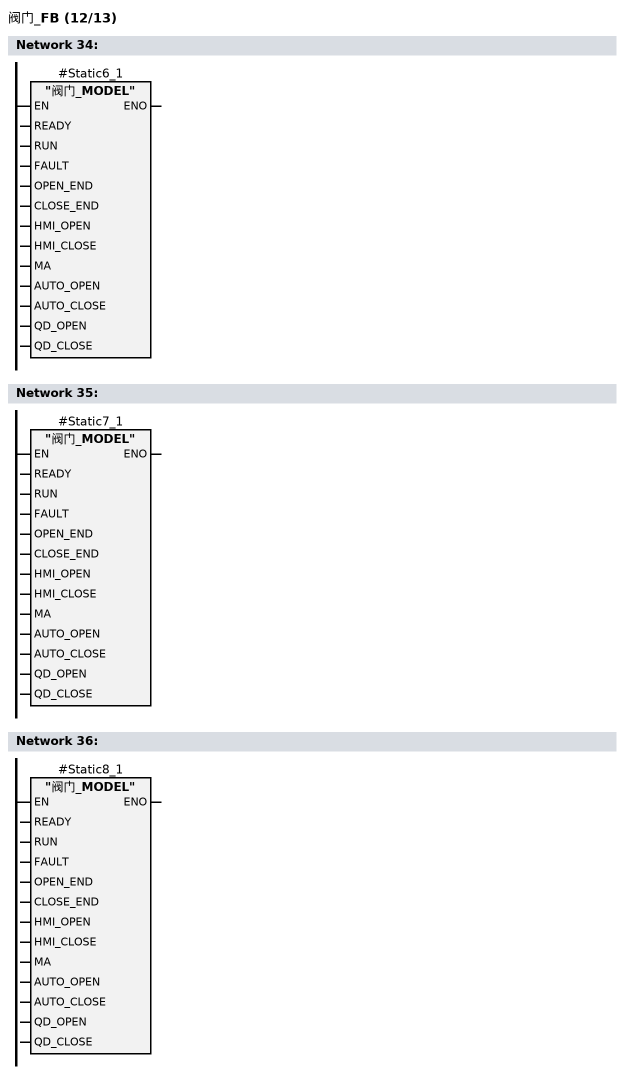
   RUNG wire#powerrail
      #Static6_1(READY :=, RUN :=, FAULT :=, OPEN_END :=, CLOSE_END :=, HMI_OPEN :=, HMI_CLOSE :=, MA :=, AUTO_OPEN :=, AUTO_CLOSE :=, QD_OPEN :=, QD_CLOSE :=)
   END_RUNG
   // the same network as SCL:
   #Static6_1();   // "阀门_MODEL"
END_REGION

REGION Network 35
   RUNG wire#powerrail
      #Static7_1(READY :=, RUN :=, FAULT :=, OPEN_END :=, CLOSE_END :=, HMI_OPEN :=, HMI_CLOSE :=, MA :=, AUTO_OPEN :=, AUTO_CLOSE :=, QD_OPEN :=, QD_CLOSE :=)
   END_RUNG
   // the same network as SCL:
   #Static7_1();   // "阀门_MODEL"
END_REGION

REGION Network 36
   RUNG wire#powerrail
      #Static8_1(READY :=, RUN :=, FAULT :=, OPEN_END :=, CLOSE_END :=, HMI_OPEN :=, HMI_CLOSE :=, MA :=, AUTO_OPEN :=, AUTO_CLOSE :=, QD_OPEN :=, QD_CLOSE :=)
   END_RUNG
   // the same network as SCL:
   #Static8_1();   // "阀门_MODEL"
END_REGION

REGION Network 37
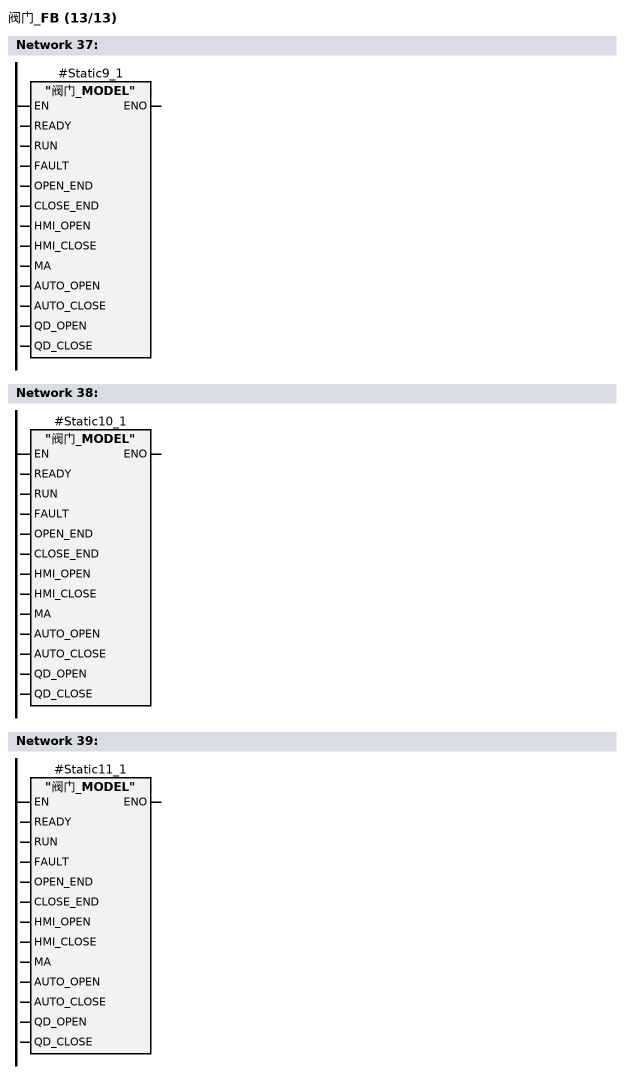
   RUNG wire#powerrail
      #Static9_1(READY :=, RUN :=, FAULT :=, OPEN_END :=, CLOSE_END :=, HMI_OPEN :=, HMI_CLOSE :=, MA :=, AUTO_OPEN :=, AUTO_CLOSE :=, QD_OPEN :=, QD_CLOSE :=)
   END_RUNG
   // the same network as SCL:
   #Static9_1();   // "阀门_MODEL"
END_REGION

REGION Network 38
   RUNG wire#powerrail
      #Static10_1(READY :=, RUN :=, FAULT :=, OPEN_END :=, CLOSE_END :=, HMI_OPEN :=, HMI_CLOSE :=, MA :=, AUTO_OPEN :=, AUTO_CLOSE :=, QD_OPEN :=, QD_CLOSE :=)
   END_RUNG
   // the same network as SCL:
   #Static10_1();   // "阀门_MODEL"
END_REGION

REGION Network 39
   RUNG wire#powerrail
      #Static11_1(READY :=, RUN :=, FAULT :=, OPEN_END :=, CLOSE_END :=, HMI_OPEN :=, HMI_CLOSE :=, MA :=, AUTO_OPEN :=, AUTO_CLOSE :=, QD_OPEN :=, QD_CLOSE :=)
   END_RUNG
   // the same network as SCL:
   #Static11_1();   // "阀门_MODEL"
END_REGION
END_FUNCTION_BLOCK

FUNCTION_BLOCK "引水阀和排气阀FB"   // FB12, LAD
{ S7_Optimized_Access := 'FALSE' }
VERSION : 0.1
   VAR
      "1#炉体循环水泵引水电磁阀" : "引水排气块";
      "1#炉体循环水泵排气电磁阀" : "引水排气块";
      "2#炉体循环水泵引水电磁阀" : "引水排气块";
      "2#炉体循环水泵排气电磁阀" : "引水排气块";
      "3#炉体循环水泵引水电磁阀" : "引水排气块";
      "3#炉体循环水泵排气电磁阀" : "引水排气块";
      "1#电极循环水泵引水电磁阀" : "引水排气块";
      "1#电极循环水泵排气电磁阀" : "引水排气块";
      "2#电极循环水泵引水电磁阀" : "引水排气块";
      "2#电极循环水泵排气电磁阀" : "引水排气块";
      "3#电极循环水泵引水电磁阀" : "引水排气块";
      "3#电极循环水泵排气电磁阀" : "引水排气块";
      "4#电极循环水泵引水电磁阀" : "引水排气块";
      "4#电极循环水泵排气电磁阀" : "引水排气块";
      "1#净环热水泵引水电磁阀" : "引水排气块";
      "1#净环热水泵排气电磁阀" : "引水排气块";
      "2#净环热水泵引水电磁阀" : "引水排气块";
      "2#净环热水泵排气电磁阀" : "引水排气块";
      "3#净环热水泵引水电磁阀" : "引水排气块";
      "3#净环热水泵排气电磁阀" : "引水排气块";
      "4#净环热水泵引水电磁阀" : "引水排气块";
      "4#净环热水泵排气电磁阀" : "引水排气块";
      "5#净环热水泵引水电磁阀" : "引水排气块";
      "5#净环热水泵排气电磁阀" : "引水排气块";
      "1#浊环热水泵引水电磁阀" : "引水排气块";
      "1#浊环热水泵排气电磁阀" : "引水排气块";
      "2#浊环热水泵引水电磁阀" : "引水排气块";
      "2#浊环热水泵排气电磁阀" : "引水排气块";
      "3#浊环热水泵引水电磁阀" : "引水排气块";
      "3#浊环热水泵排气电磁阀" : "引水排气块";
      "4#浊环热水泵引水电磁阀" : "引水排气块";
      "4#浊环热水泵排气电磁阀" : "引水排气块";
      "5#浊环热水泵引水电磁阀" : "引水排气块";
      "5#浊环热水泵排气电磁阀" : "引水排气块";
      "6#浊环热水泵引水电磁阀" : "引水排气块";
      "6#浊环热水泵排气电磁阀" : "引水排气块";
      "7#浊环热水泵引水电磁阀" : "引水排气块";
      "7#浊环热水泵排气电磁阀" : "引水排气块";
      "8#浊环热水泵引水电磁阀" : "引水排气块";
      "8#浊环热水泵排气电磁阀" : "引水排气块";
      "1#冲渣泵引水电磁阀" : "引水排气块";
      "1#冲渣泵排气电磁阀" : "引水排气块";
      "2#冲渣泵引水电磁阀" : "引水排气块";
      "2#冲渣泵排气电磁阀" : "引水排气块";
      "3#冲渣泵引水电磁阀" : "引水排气块";
      "3#冲渣泵排气电磁阀" : "引水排气块";
      "4#冲渣泵引水电磁阀" : "引水排气块";
      "4#冲渣泵排气电磁阀" : "引水排气块";
      "5#冲渣泵引水电磁阀" : "引水排气块";
      "5#冲渣泵排气电磁阀" : "引水排气块";
      "6#冲渣泵引水电磁阀" : "引水排气块";
      "6#冲渣泵排气电磁阀" : "引水排气块";
      "7#冲渣泵引水电磁阀" : "引水排气块";
      "7#冲渣泵排气电磁阀" : "引水排气块";
      "8#冲渣泵引水电磁阀" : "引水排气块";
      "8#冲渣泵排气电磁阀" : "引水排气块";
      "1#柴油泵引水电磁阀" : "引水排气块";
      "1#柴油泵排气电磁阀" : "引水排气块";
      "2#柴油泵引水电磁阀" : "引水排气块";
      "2#柴油泵排气电磁阀" : "引水排气块";
      "1#炉冲渣报警" : "引水排气块";
      "2#炉冲渣报警" : "引水排气块";
      窑冷却泵引水电池阀 : "引水排气块";
      窑冷却泵排气电池阀 : "引水排气块";
      Static9 : "引水排气块";
      Static10 : "引水排气块";
      Static11 : "引水排气块";
      Static12 : "引水排气块";
      Static13 : "引水排气块";
      Static14 : "引水排气块";
      Static15 : "引水排气块";
      Static16 : "引水排气块";
      Static17 : "引水排气块";
      Static18 : "引水排气块";
      Static19 : "引水排气块";
      Static20 : "引水排气块";
      Static21 : "引水排气块";
      Static22 : "引水排气块";
      Static23 : "引水排气块";
      Static24 : "引水排气块";
      Static25 : "引水排气块";
      Static26 : "引水排气块";
      Static27 : "引水排气块";
      Static28 : "引水排气块";
      Static29 : "引水排气块";
      Static30 : "引水排气块";
      Static31 : "引水排气块";
      Static32 : "引水排气块";
      Static33 : "引水排气块";
      Static34 : "引水排气块";
      Static35 : "引水排气块";
      Static36 : "引水排气块";
   END_VAR
BEGIN

REGION Network 1
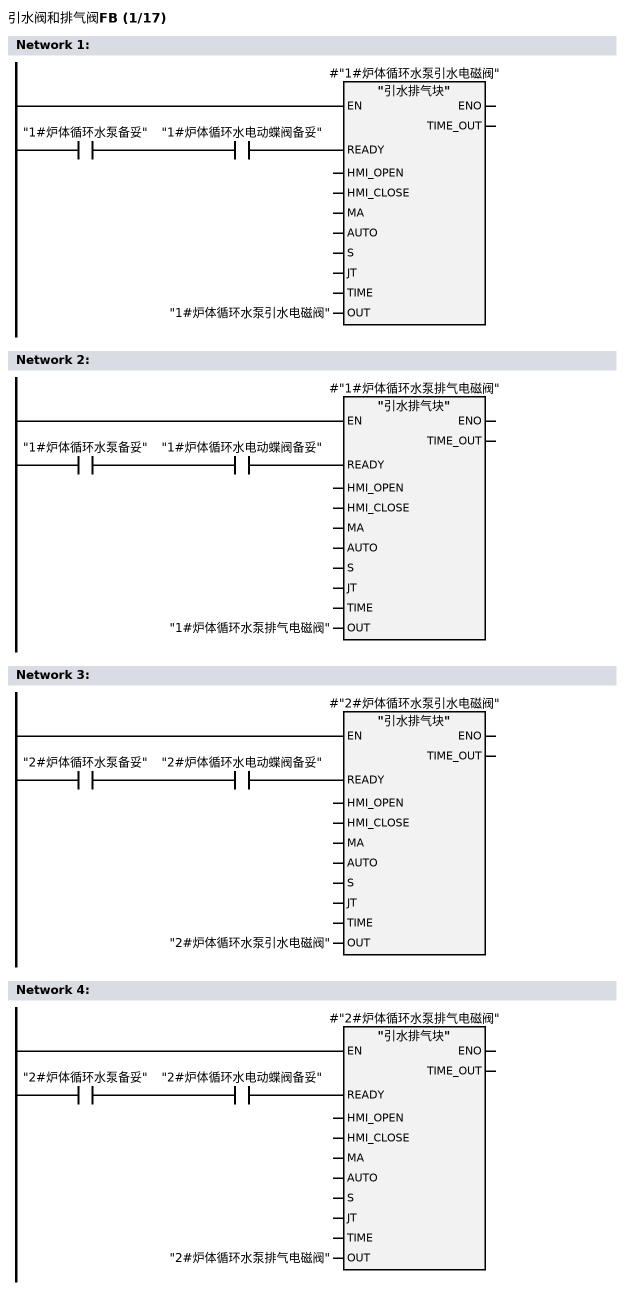
   RUNG wire#powerrail
      #"1#炉体循环水泵引水电磁阀"(READY := wire#w1, HMI_OPEN :=, HMI_CLOSE :=, MA :=, AUTO :=, S :=, JT :=, "TIME" :=, OUT := "1#炉体循环水泵引水电磁阀", TIME_OUT =>)
   END_RUNG
   RUNG wire#powerrail
      Contact( "1#炉体循环水泵备妥" )
      Contact( "1#炉体循环水电动蝶阀备妥" )
   END_RUNG wire#w1
   // the same network as SCL:
   #"1#炉体循环水泵引水电磁阀"(READY := "1#炉体循环水泵备妥" AND "1#炉体循环水电动蝶阀备妥", OUT := "1#炉体循环水泵引水电磁阀");   // "引水排气块"
END_REGION

REGION Network 2
   RUNG wire#powerrail
      #"1#炉体循环水泵排气电磁阀"(READY := wire#w1, HMI_OPEN :=, HMI_CLOSE :=, MA :=, AUTO :=, S :=, JT :=, "TIME" :=, OUT := "1#炉体循环水泵排气电磁阀", TIME_OUT =>)
   END_RUNG
   RUNG wire#powerrail
      Contact( "1#炉体循环水泵备妥" )
      Contact( "1#炉体循环水电动蝶阀备妥" )
   END_RUNG wire#w1
   // the same network as SCL:
   #"1#炉体循环水泵排气电磁阀"(READY := "1#炉体循环水泵备妥" AND "1#炉体循环水电动蝶阀备妥", OUT := "1#炉体循环水泵排气电磁阀");   // "引水排气块"
END_REGION

REGION Network 3
   RUNG wire#powerrail
      #"2#炉体循环水泵引水电磁阀"(READY := wire#w1, HMI_OPEN :=, HMI_CLOSE :=, MA :=, AUTO :=, S :=, JT :=, "TIME" :=, OUT := "2#炉体循环水泵引水电磁阀", TIME_OUT =>)
   END_RUNG
   RUNG wire#powerrail
      Contact( "2#炉体循环水泵备妥" )
      Contact( "2#炉体循环水电动蝶阀备妥" )
   END_RUNG wire#w1
   // the same network as SCL:
   #"2#炉体循环水泵引水电磁阀"(READY := "2#炉体循环水泵备妥" AND "2#炉体循环水电动蝶阀备妥", OUT := "2#炉体循环水泵引水电磁阀");   // "引水排气块"
END_REGION

REGION Network 4
   RUNG wire#powerrail
      #"2#炉体循环水泵排气电磁阀"(READY := wire#w1, HMI_OPEN :=, HMI_CLOSE :=, MA :=, AUTO :=, S :=, JT :=, "TIME" :=, OUT := "2#炉体循环水泵排气电磁阀", TIME_OUT =>)
   END_RUNG
   RUNG wire#powerrail
      Contact( "2#炉体循环水泵备妥" )
      Contact( "2#炉体循环水电动蝶阀备妥" )
   END_RUNG wire#w1
   // the same network as SCL:
   #"2#炉体循环水泵排气电磁阀"(READY := "2#炉体循环水泵备妥" AND "2#炉体循环水电动蝶阀备妥", OUT := "2#炉体循环水泵排气电磁阀");   // "引水排气块"
END_REGION

REGION Network 5
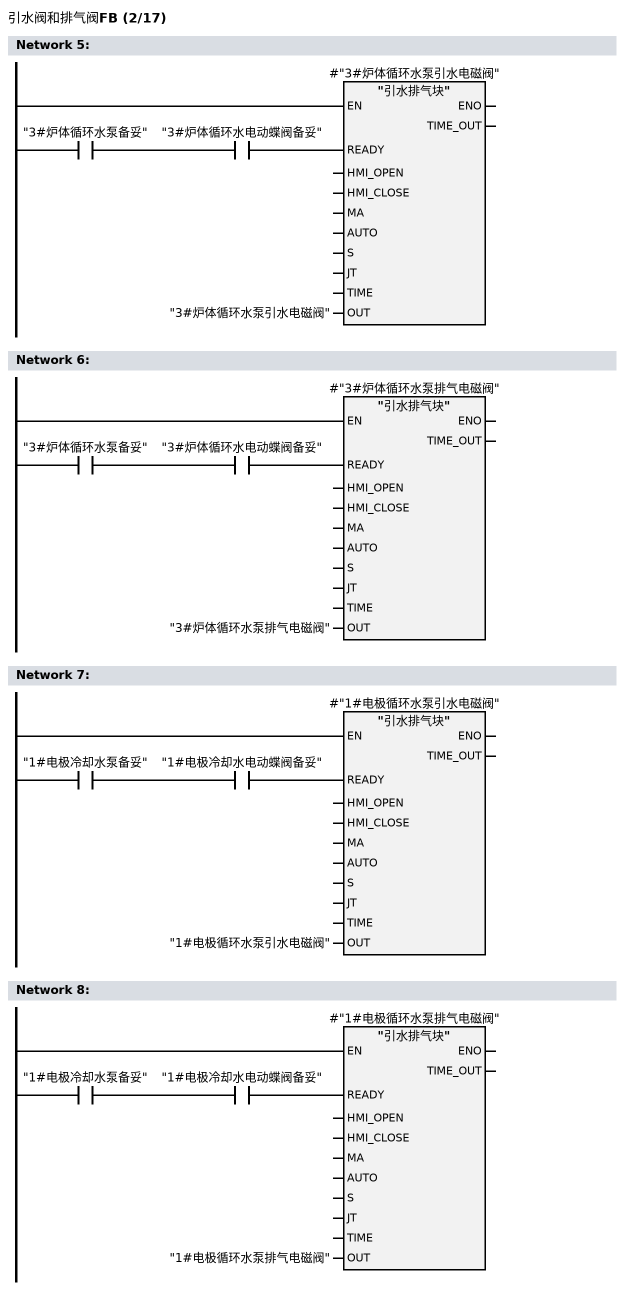
   RUNG wire#powerrail
      #"3#炉体循环水泵引水电磁阀"(READY := wire#w1, HMI_OPEN :=, HMI_CLOSE :=, MA :=, AUTO :=, S :=, JT :=, "TIME" :=, OUT := "3#炉体循环水泵引水电磁阀", TIME_OUT =>)
   END_RUNG
   RUNG wire#powerrail
      Contact( "3#炉体循环水泵备妥" )
      Contact( "3#炉体循环水电动蝶阀备妥" )
   END_RUNG wire#w1
   // the same network as SCL:
   #"3#炉体循环水泵引水电磁阀"(READY := "3#炉体循环水泵备妥" AND "3#炉体循环水电动蝶阀备妥", OUT := "3#炉体循环水泵引水电磁阀");   // "引水排气块"
END_REGION

REGION Network 6
   RUNG wire#powerrail
      #"3#炉体循环水泵排气电磁阀"(READY := wire#w1, HMI_OPEN :=, HMI_CLOSE :=, MA :=, AUTO :=, S :=, JT :=, "TIME" :=, OUT := "3#炉体循环水泵排气电磁阀", TIME_OUT =>)
   END_RUNG
   RUNG wire#powerrail
      Contact( "3#炉体循环水泵备妥" )
      Contact( "3#炉体循环水电动蝶阀备妥" )
   END_RUNG wire#w1
   // the same network as SCL:
   #"3#炉体循环水泵排气电磁阀"(READY := "3#炉体循环水泵备妥" AND "3#炉体循环水电动蝶阀备妥", OUT := "3#炉体循环水泵排气电磁阀");   // "引水排气块"
END_REGION

REGION Network 7
   RUNG wire#powerrail
      #"1#电极循环水泵引水电磁阀"(READY := wire#w1, HMI_OPEN :=, HMI_CLOSE :=, MA :=, AUTO :=, S :=, JT :=, "TIME" :=, OUT := "1#电极循环水泵引水电磁阀", TIME_OUT =>)
   END_RUNG
   RUNG wire#powerrail
      Contact( "1#电极冷却水泵备妥" )
      Contact( "1#电极冷却水电动蝶阀备妥" )
   END_RUNG wire#w1
   // the same network as SCL:
   #"1#电极循环水泵引水电磁阀"(READY := "1#电极冷却水泵备妥" AND "1#电极冷却水电动蝶阀备妥", OUT := "1#电极循环水泵引水电磁阀");   // "引水排气块"
END_REGION

REGION Network 8
   RUNG wire#powerrail
      #"1#电极循环水泵排气电磁阀"(READY := wire#w1, HMI_OPEN :=, HMI_CLOSE :=, MA :=, AUTO :=, S :=, JT :=, "TIME" :=, OUT := "1#电极循环水泵排气电磁阀", TIME_OUT =>)
   END_RUNG
   RUNG wire#powerrail
      Contact( "1#电极冷却水泵备妥" )
      Contact( "1#电极冷却水电动蝶阀备妥" )
   END_RUNG wire#w1
   // the same network as SCL:
   #"1#电极循环水泵排气电磁阀"(READY := "1#电极冷却水泵备妥" AND "1#电极冷却水电动蝶阀备妥", OUT := "1#电极循环水泵排气电磁阀");   // "引水排气块"
END_REGION

REGION Network 9
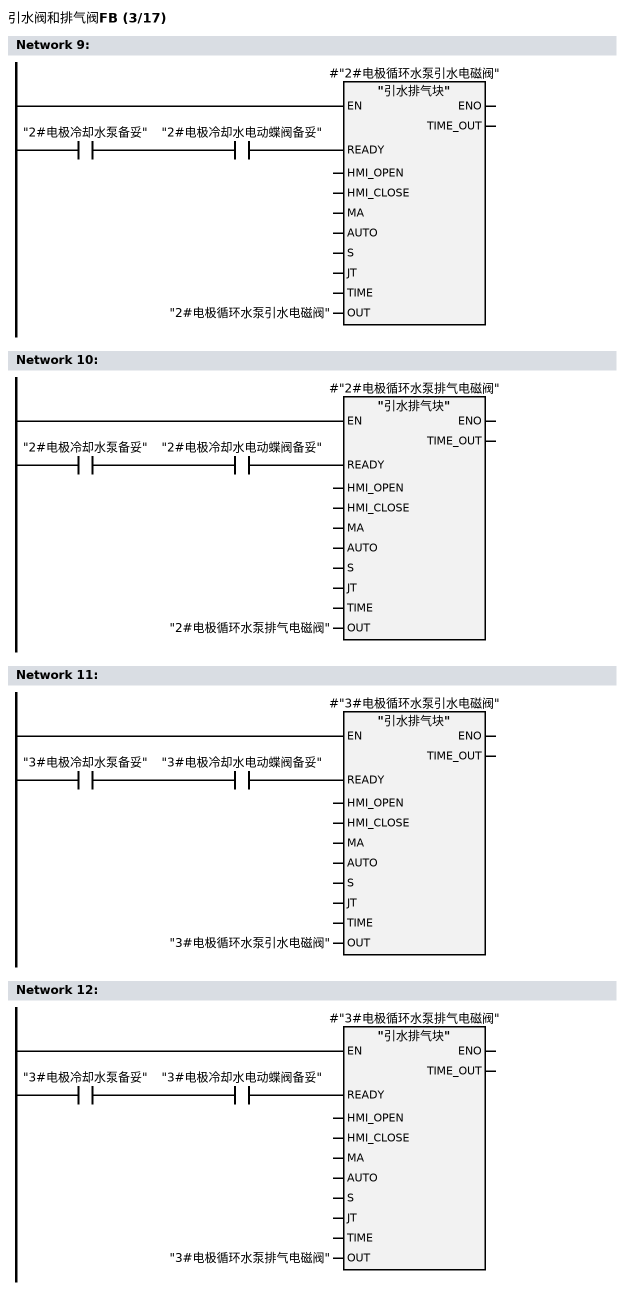
   RUNG wire#powerrail
      #"2#电极循环水泵引水电磁阀"(READY := wire#w1, HMI_OPEN :=, HMI_CLOSE :=, MA :=, AUTO :=, S :=, JT :=, "TIME" :=, OUT := "2#电极循环水泵引水电磁阀", TIME_OUT =>)
   END_RUNG
   RUNG wire#powerrail
      Contact( "2#电极冷却水泵备妥" )
      Contact( "2#电极冷却水电动蝶阀备妥" )
   END_RUNG wire#w1
   // the same network as SCL:
   #"2#电极循环水泵引水电磁阀"(READY := "2#电极冷却水泵备妥" AND "2#电极冷却水电动蝶阀备妥", OUT := "2#电极循环水泵引水电磁阀");   // "引水排气块"
END_REGION

REGION Network 10
   RUNG wire#powerrail
      #"2#电极循环水泵排气电磁阀"(READY := wire#w1, HMI_OPEN :=, HMI_CLOSE :=, MA :=, AUTO :=, S :=, JT :=, "TIME" :=, OUT := "2#电极循环水泵排气电磁阀", TIME_OUT =>)
   END_RUNG
   RUNG wire#powerrail
      Contact( "2#电极冷却水泵备妥" )
      Contact( "2#电极冷却水电动蝶阀备妥" )
   END_RUNG wire#w1
   // the same network as SCL:
   #"2#电极循环水泵排气电磁阀"(READY := "2#电极冷却水泵备妥" AND "2#电极冷却水电动蝶阀备妥", OUT := "2#电极循环水泵排气电磁阀");   // "引水排气块"
END_REGION

REGION Network 11
   RUNG wire#powerrail
      #"3#电极循环水泵引水电磁阀"(READY := wire#w1, HMI_OPEN :=, HMI_CLOSE :=, MA :=, AUTO :=, S :=, JT :=, "TIME" :=, OUT := "3#电极循环水泵引水电磁阀", TIME_OUT =>)
   END_RUNG
   RUNG wire#powerrail
      Contact( "3#电极冷却水泵备妥" )
      Contact( "3#电极冷却水电动蝶阀备妥" )
   END_RUNG wire#w1
   // the same network as SCL:
   #"3#电极循环水泵引水电磁阀"(READY := "3#电极冷却水泵备妥" AND "3#电极冷却水电动蝶阀备妥", OUT := "3#电极循环水泵引水电磁阀");   // "引水排气块"
END_REGION

REGION Network 12
   RUNG wire#powerrail
      #"3#电极循环水泵排气电磁阀"(READY := wire#w1, HMI_OPEN :=, HMI_CLOSE :=, MA :=, AUTO :=, S :=, JT :=, "TIME" :=, OUT := "3#电极循环水泵排气电磁阀", TIME_OUT =>)
   END_RUNG
   RUNG wire#powerrail
      Contact( "3#电极冷却水泵备妥" )
      Contact( "3#电极冷却水电动蝶阀备妥" )
   END_RUNG wire#w1
   // the same network as SCL:
   #"3#电极循环水泵排气电磁阀"(READY := "3#电极冷却水泵备妥" AND "3#电极冷却水电动蝶阀备妥", OUT := "3#电极循环水泵排气电磁阀");   // "引水排气块"
END_REGION

REGION Network 13
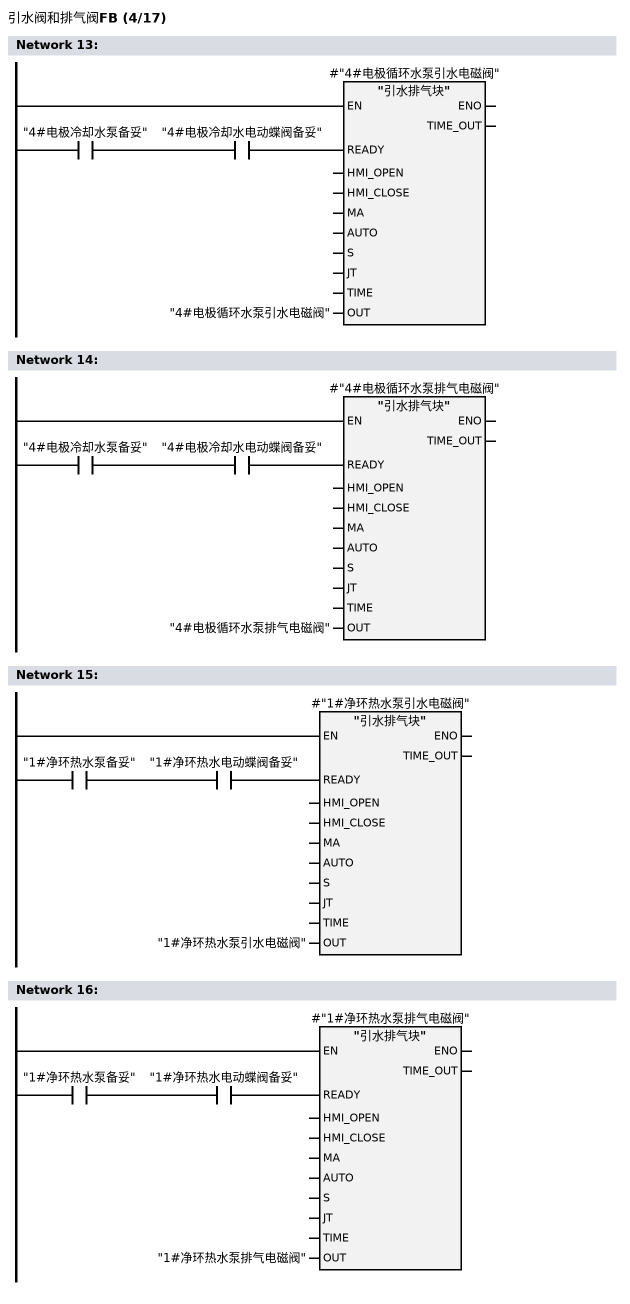
   RUNG wire#powerrail
      #"4#电极循环水泵引水电磁阀"(READY := wire#w1, HMI_OPEN :=, HMI_CLOSE :=, MA :=, AUTO :=, S :=, JT :=, "TIME" :=, OUT := "4#电极循环水泵引水电磁阀", TIME_OUT =>)
   END_RUNG
   RUNG wire#powerrail
      Contact( "4#电极冷却水泵备妥" )
      Contact( "4#电极冷却水电动蝶阀备妥" )
   END_RUNG wire#w1
   // the same network as SCL:
   #"4#电极循环水泵引水电磁阀"(READY := "4#电极冷却水泵备妥" AND "4#电极冷却水电动蝶阀备妥", OUT := "4#电极循环水泵引水电磁阀");   // "引水排气块"
END_REGION

REGION Network 14
   RUNG wire#powerrail
      #"4#电极循环水泵排气电磁阀"(READY := wire#w1, HMI_OPEN :=, HMI_CLOSE :=, MA :=, AUTO :=, S :=, JT :=, "TIME" :=, OUT := "4#电极循环水泵排气电磁阀", TIME_OUT =>)
   END_RUNG
   RUNG wire#powerrail
      Contact( "4#电极冷却水泵备妥" )
      Contact( "4#电极冷却水电动蝶阀备妥" )
   END_RUNG wire#w1
   // the same network as SCL:
   #"4#电极循环水泵排气电磁阀"(READY := "4#电极冷却水泵备妥" AND "4#电极冷却水电动蝶阀备妥", OUT := "4#电极循环水泵排气电磁阀");   // "引水排气块"
END_REGION

REGION Network 15
   RUNG wire#powerrail
      #"1#净环热水泵引水电磁阀"(READY := wire#w1, HMI_OPEN :=, HMI_CLOSE :=, MA :=, AUTO :=, S :=, JT :=, "TIME" :=, OUT := "1#净环热水泵引水电磁阀", TIME_OUT =>)
   END_RUNG
   RUNG wire#powerrail
      Contact( "1#净环热水泵备妥" )
      Contact( "1#净环热水电动蝶阀备妥" )
   END_RUNG wire#w1
   // the same network as SCL:
   #"1#净环热水泵引水电磁阀"(READY := "1#净环热水泵备妥" AND "1#净环热水电动蝶阀备妥", OUT := "1#净环热水泵引水电磁阀");   // "引水排气块"
END_REGION

REGION Network 16
   RUNG wire#powerrail
      #"1#净环热水泵排气电磁阀"(READY := wire#w1, HMI_OPEN :=, HMI_CLOSE :=, MA :=, AUTO :=, S :=, JT :=, "TIME" :=, OUT := "1#净环热水泵排气电磁阀", TIME_OUT =>)
   END_RUNG
   RUNG wire#powerrail
      Contact( "1#净环热水泵备妥" )
      Contact( "1#净环热水电动蝶阀备妥" )
   END_RUNG wire#w1
   // the same network as SCL:
   #"1#净环热水泵排气电磁阀"(READY := "1#净环热水泵备妥" AND "1#净环热水电动蝶阀备妥", OUT := "1#净环热水泵排气电磁阀");   // "引水排气块"
END_REGION

REGION Network 17
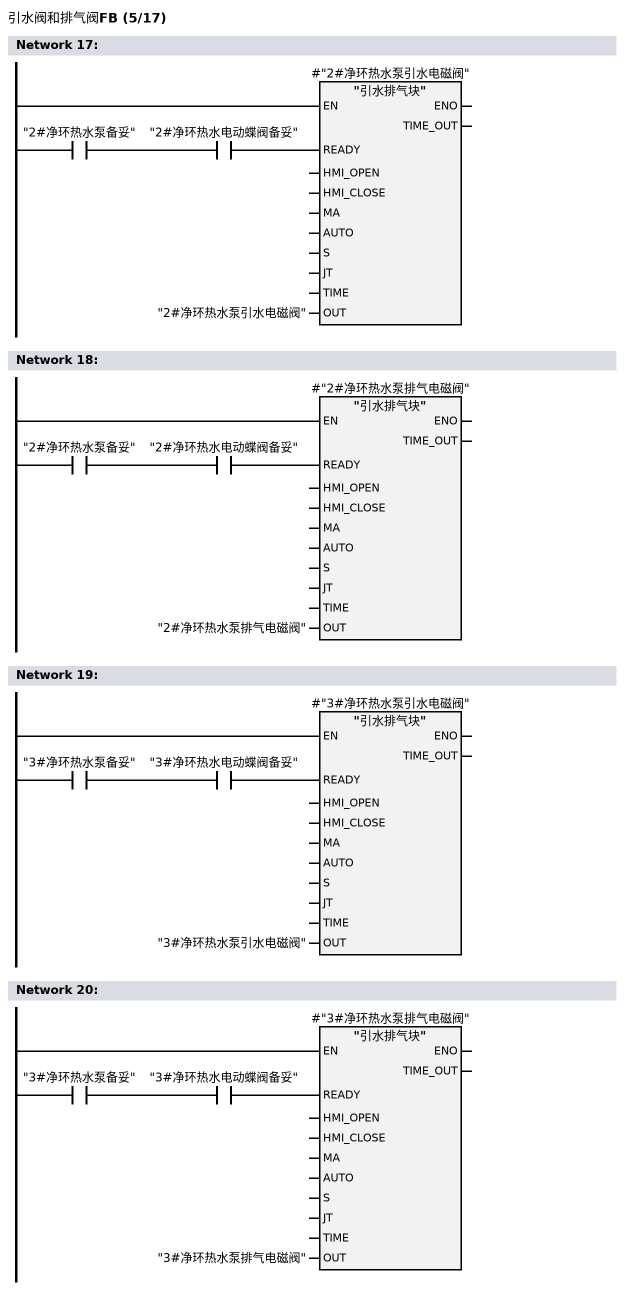
   RUNG wire#powerrail
      #"2#净环热水泵引水电磁阀"(READY := wire#w1, HMI_OPEN :=, HMI_CLOSE :=, MA :=, AUTO :=, S :=, JT :=, "TIME" :=, OUT := "2#净环热水泵引水电磁阀", TIME_OUT =>)
   END_RUNG
   RUNG wire#powerrail
      Contact( "2#净环热水泵备妥" )
      Contact( "2#净环热水电动蝶阀备妥" )
   END_RUNG wire#w1
   // the same network as SCL:
   #"2#净环热水泵引水电磁阀"(READY := "2#净环热水泵备妥" AND "2#净环热水电动蝶阀备妥", OUT := "2#净环热水泵引水电磁阀");   // "引水排气块"
END_REGION

REGION Network 18
   RUNG wire#powerrail
      #"2#净环热水泵排气电磁阀"(READY := wire#w1, HMI_OPEN :=, HMI_CLOSE :=, MA :=, AUTO :=, S :=, JT :=, "TIME" :=, OUT := "2#净环热水泵排气电磁阀", TIME_OUT =>)
   END_RUNG
   RUNG wire#powerrail
      Contact( "2#净环热水泵备妥" )
      Contact( "2#净环热水电动蝶阀备妥" )
   END_RUNG wire#w1
   // the same network as SCL:
   #"2#净环热水泵排气电磁阀"(READY := "2#净环热水泵备妥" AND "2#净环热水电动蝶阀备妥", OUT := "2#净环热水泵排气电磁阀");   // "引水排气块"
END_REGION

REGION Network 19
   RUNG wire#powerrail
      #"3#净环热水泵引水电磁阀"(READY := wire#w1, HMI_OPEN :=, HMI_CLOSE :=, MA :=, AUTO :=, S :=, JT :=, "TIME" :=, OUT := "3#净环热水泵引水电磁阀", TIME_OUT =>)
   END_RUNG
   RUNG wire#powerrail
      Contact( "3#净环热水泵备妥" )
      Contact( "3#净环热水电动蝶阀备妥" )
   END_RUNG wire#w1
   // the same network as SCL:
   #"3#净环热水泵引水电磁阀"(READY := "3#净环热水泵备妥" AND "3#净环热水电动蝶阀备妥", OUT := "3#净环热水泵引水电磁阀");   // "引水排气块"
END_REGION

REGION Network 20
   RUNG wire#powerrail
      #"3#净环热水泵排气电磁阀"(READY := wire#w1, HMI_OPEN :=, HMI_CLOSE :=, MA :=, AUTO :=, S :=, JT :=, "TIME" :=, OUT := "3#净环热水泵排气电磁阀", TIME_OUT =>)
   END_RUNG
   RUNG wire#powerrail
      Contact( "3#净环热水泵备妥" )
      Contact( "3#净环热水电动蝶阀备妥" )
   END_RUNG wire#w1
   // the same network as SCL:
   #"3#净环热水泵排气电磁阀"(READY := "3#净环热水泵备妥" AND "3#净环热水电动蝶阀备妥", OUT := "3#净环热水泵排气电磁阀");   // "引水排气块"
END_REGION

REGION Network 21
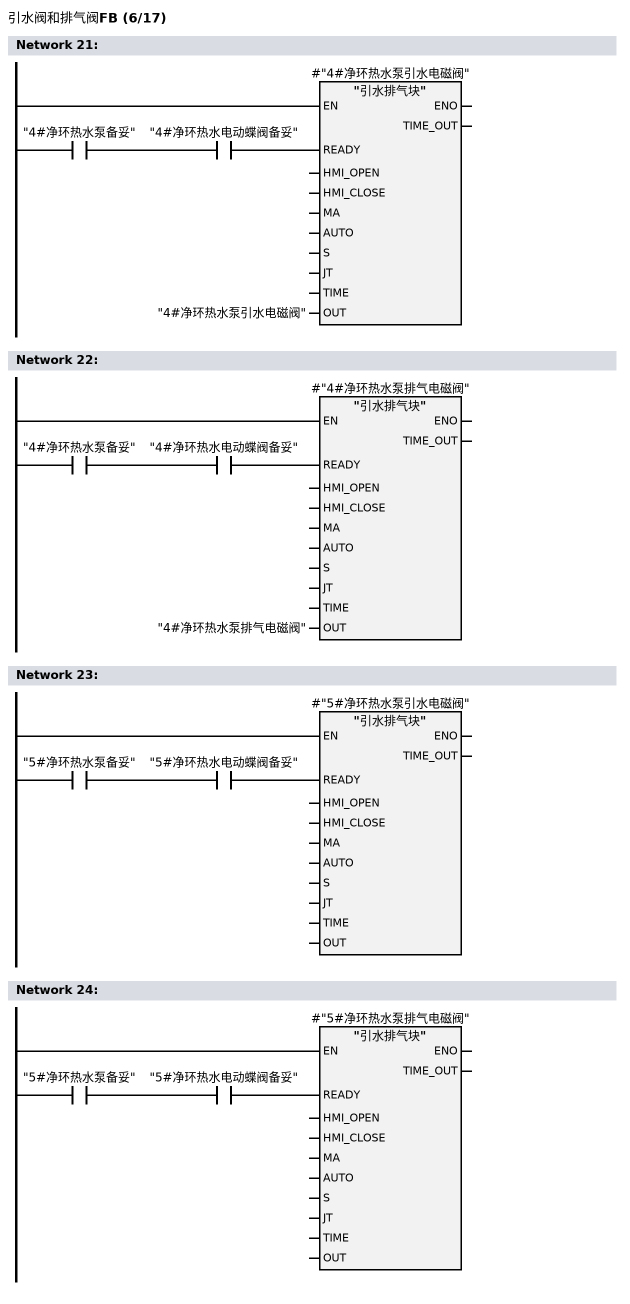
   RUNG wire#powerrail
      #"4#净环热水泵引水电磁阀"(READY := wire#w1, HMI_OPEN :=, HMI_CLOSE :=, MA :=, AUTO :=, S :=, JT :=, "TIME" :=, OUT := "4#净环热水泵引水电磁阀", TIME_OUT =>)
   END_RUNG
   RUNG wire#powerrail
      Contact( "4#净环热水泵备妥" )
      Contact( "4#净环热水电动蝶阀备妥" )
   END_RUNG wire#w1
   // the same network as SCL:
   #"4#净环热水泵引水电磁阀"(READY := "4#净环热水泵备妥" AND "4#净环热水电动蝶阀备妥", OUT := "4#净环热水泵引水电磁阀");   // "引水排气块"
END_REGION

REGION Network 22
   RUNG wire#powerrail
      #"4#净环热水泵排气电磁阀"(READY := wire#w1, HMI_OPEN :=, HMI_CLOSE :=, MA :=, AUTO :=, S :=, JT :=, "TIME" :=, OUT := "4#净环热水泵排气电磁阀", TIME_OUT =>)
   END_RUNG
   RUNG wire#powerrail
      Contact( "4#净环热水泵备妥" )
      Contact( "4#净环热水电动蝶阀备妥" )
   END_RUNG wire#w1
   // the same network as SCL:
   #"4#净环热水泵排气电磁阀"(READY := "4#净环热水泵备妥" AND "4#净环热水电动蝶阀备妥", OUT := "4#净环热水泵排气电磁阀");   // "引水排气块"
END_REGION

REGION Network 23
   RUNG wire#powerrail
      #"5#净环热水泵引水电磁阀"(READY := wire#w1, HMI_OPEN :=, HMI_CLOSE :=, MA :=, AUTO :=, S :=, JT :=, "TIME" :=, OUT :=, TIME_OUT =>)
   END_RUNG
   RUNG wire#powerrail
      Contact( "5#净环热水泵备妥" )
      Contact( "5#净环热水电动蝶阀备妥" )
   END_RUNG wire#w1
   // the same network as SCL:
   #"5#净环热水泵引水电磁阀"(READY := "5#净环热水泵备妥" AND "5#净环热水电动蝶阀备妥");   // "引水排气块"
END_REGION

REGION Network 24
   RUNG wire#powerrail
      #"5#净环热水泵排气电磁阀"(READY := wire#w1, HMI_OPEN :=, HMI_CLOSE :=, MA :=, AUTO :=, S :=, JT :=, "TIME" :=, OUT :=, TIME_OUT =>)
   END_RUNG
   RUNG wire#powerrail
      Contact( "5#净环热水泵备妥" )
      Contact( "5#净环热水电动蝶阀备妥" )
   END_RUNG wire#w1
   // the same network as SCL:
   #"5#净环热水泵排气电磁阀"(READY := "5#净环热水泵备妥" AND "5#净环热水电动蝶阀备妥");   // "引水排气块"
END_REGION

REGION Network 25
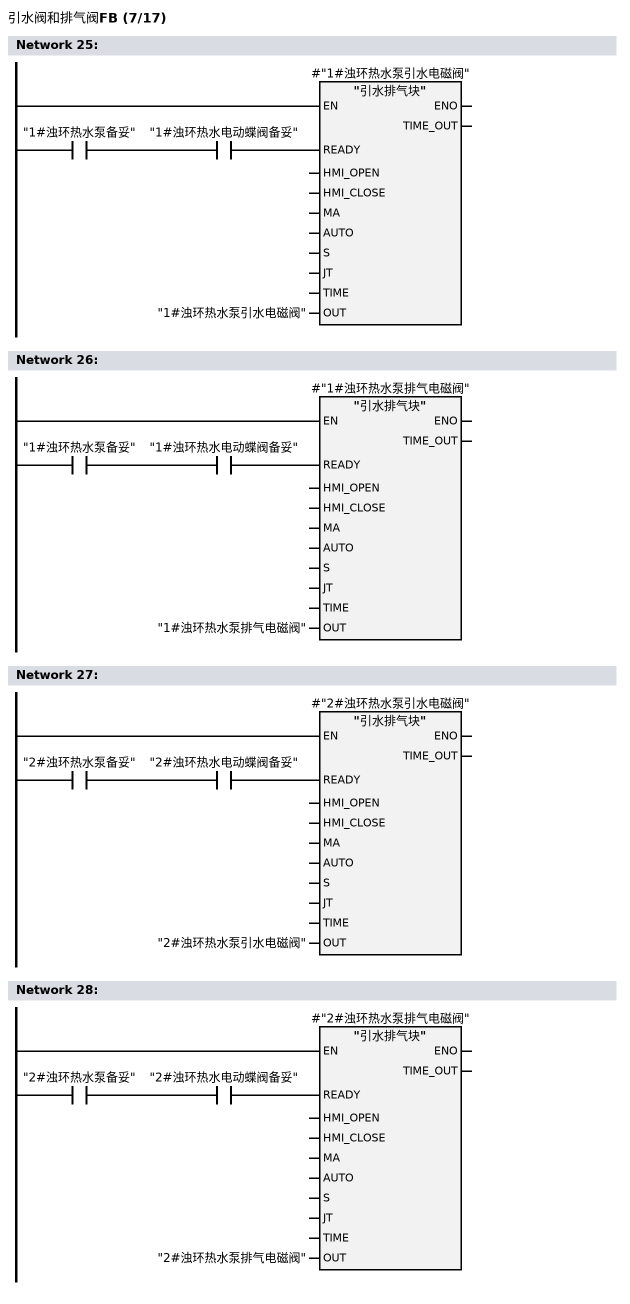
   RUNG wire#powerrail
      #"1#浊环热水泵引水电磁阀"(READY := wire#w1, HMI_OPEN :=, HMI_CLOSE :=, MA :=, AUTO :=, S :=, JT :=, "TIME" :=, OUT := "1#浊环热水泵引水电磁阀", TIME_OUT =>)
   END_RUNG
   RUNG wire#powerrail
      Contact( "1#浊环热水泵备妥" )
      Contact( "1#浊环热水电动蝶阀备妥" )
   END_RUNG wire#w1
   // the same network as SCL:
   #"1#浊环热水泵引水电磁阀"(READY := "1#浊环热水泵备妥" AND "1#浊环热水电动蝶阀备妥", OUT := "1#浊环热水泵引水电磁阀");   // "引水排气块"
END_REGION

REGION Network 26
   RUNG wire#powerrail
      #"1#浊环热水泵排气电磁阀"(READY := wire#w1, HMI_OPEN :=, HMI_CLOSE :=, MA :=, AUTO :=, S :=, JT :=, "TIME" :=, OUT := "1#浊环热水泵排气电磁阀", TIME_OUT =>)
   END_RUNG
   RUNG wire#powerrail
      Contact( "1#浊环热水泵备妥" )
      Contact( "1#浊环热水电动蝶阀备妥" )
   END_RUNG wire#w1
   // the same network as SCL:
   #"1#浊环热水泵排气电磁阀"(READY := "1#浊环热水泵备妥" AND "1#浊环热水电动蝶阀备妥", OUT := "1#浊环热水泵排气电磁阀");   // "引水排气块"
END_REGION

REGION Network 27
   RUNG wire#powerrail
      #"2#浊环热水泵引水电磁阀"(READY := wire#w1, HMI_OPEN :=, HMI_CLOSE :=, MA :=, AUTO :=, S :=, JT :=, "TIME" :=, OUT := "2#浊环热水泵引水电磁阀", TIME_OUT =>)
   END_RUNG
   RUNG wire#powerrail
      Contact( "2#浊环热水泵备妥" )
      Contact( "2#浊环热水电动蝶阀备妥" )
   END_RUNG wire#w1
   // the same network as SCL:
   #"2#浊环热水泵引水电磁阀"(READY := "2#浊环热水泵备妥" AND "2#浊环热水电动蝶阀备妥", OUT := "2#浊环热水泵引水电磁阀");   // "引水排气块"
END_REGION

REGION Network 28
   RUNG wire#powerrail
      #"2#浊环热水泵排气电磁阀"(READY := wire#w1, HMI_OPEN :=, HMI_CLOSE :=, MA :=, AUTO :=, S :=, JT :=, "TIME" :=, OUT := "2#浊环热水泵排气电磁阀", TIME_OUT =>)
   END_RUNG
   RUNG wire#powerrail
      Contact( "2#浊环热水泵备妥" )
      Contact( "2#浊环热水电动蝶阀备妥" )
   END_RUNG wire#w1
   // the same network as SCL:
   #"2#浊环热水泵排气电磁阀"(READY := "2#浊环热水泵备妥" AND "2#浊环热水电动蝶阀备妥", OUT := "2#浊环热水泵排气电磁阀");   // "引水排气块"
END_REGION

REGION Network 29
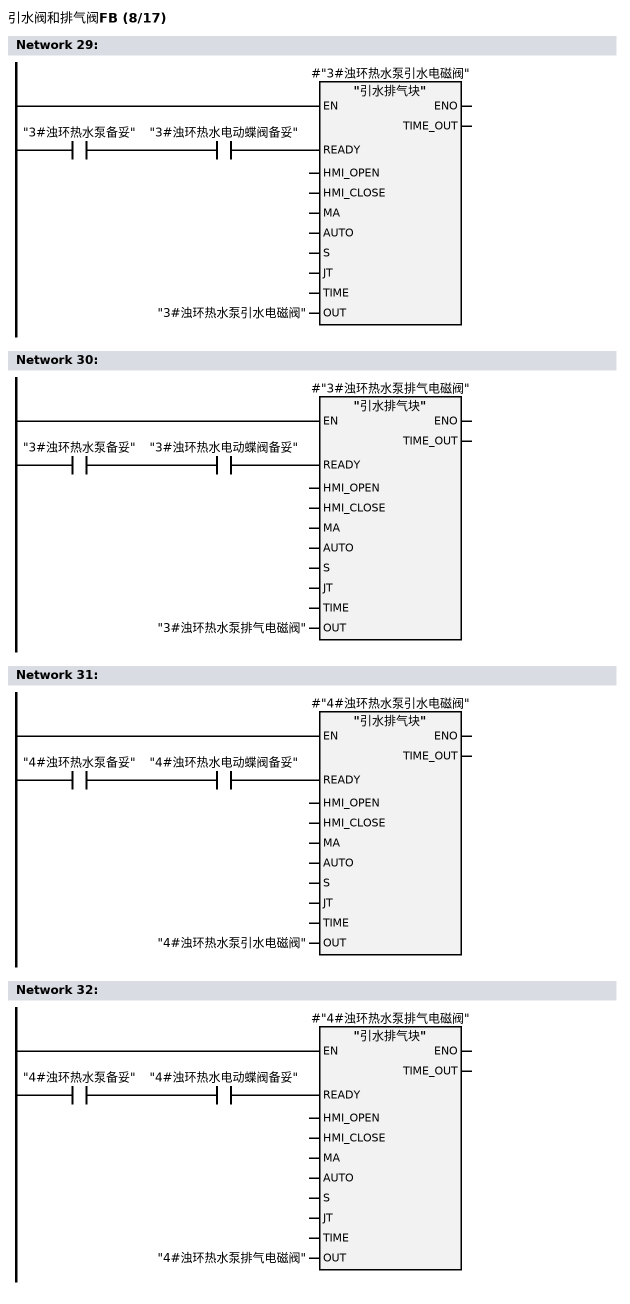
   RUNG wire#powerrail
      #"3#浊环热水泵引水电磁阀"(READY := wire#w1, HMI_OPEN :=, HMI_CLOSE :=, MA :=, AUTO :=, S :=, JT :=, "TIME" :=, OUT := "3#浊环热水泵引水电磁阀", TIME_OUT =>)
   END_RUNG
   RUNG wire#powerrail
      Contact( "3#浊环热水泵备妥" )
      Contact( "3#浊环热水电动蝶阀备妥" )
   END_RUNG wire#w1
   // the same network as SCL:
   #"3#浊环热水泵引水电磁阀"(READY := "3#浊环热水泵备妥" AND "3#浊环热水电动蝶阀备妥", OUT := "3#浊环热水泵引水电磁阀");   // "引水排气块"
END_REGION

REGION Network 30
   RUNG wire#powerrail
      #"3#浊环热水泵排气电磁阀"(READY := wire#w1, HMI_OPEN :=, HMI_CLOSE :=, MA :=, AUTO :=, S :=, JT :=, "TIME" :=, OUT := "3#浊环热水泵排气电磁阀", TIME_OUT =>)
   END_RUNG
   RUNG wire#powerrail
      Contact( "3#浊环热水泵备妥" )
      Contact( "3#浊环热水电动蝶阀备妥" )
   END_RUNG wire#w1
   // the same network as SCL:
   #"3#浊环热水泵排气电磁阀"(READY := "3#浊环热水泵备妥" AND "3#浊环热水电动蝶阀备妥", OUT := "3#浊环热水泵排气电磁阀");   // "引水排气块"
END_REGION

REGION Network 31
   RUNG wire#powerrail
      #"4#浊环热水泵引水电磁阀"(READY := wire#w1, HMI_OPEN :=, HMI_CLOSE :=, MA :=, AUTO :=, S :=, JT :=, "TIME" :=, OUT := "4#浊环热水泵引水电磁阀", TIME_OUT =>)
   END_RUNG
   RUNG wire#powerrail
      Contact( "4#浊环热水泵备妥" )
      Contact( "4#浊环热水电动蝶阀备妥" )
   END_RUNG wire#w1
   // the same network as SCL:
   #"4#浊环热水泵引水电磁阀"(READY := "4#浊环热水泵备妥" AND "4#浊环热水电动蝶阀备妥", OUT := "4#浊环热水泵引水电磁阀");   // "引水排气块"
END_REGION

REGION Network 32
   RUNG wire#powerrail
      #"4#浊环热水泵排气电磁阀"(READY := wire#w1, HMI_OPEN :=, HMI_CLOSE :=, MA :=, AUTO :=, S :=, JT :=, "TIME" :=, OUT := "4#浊环热水泵排气电磁阀", TIME_OUT =>)
   END_RUNG
   RUNG wire#powerrail
      Contact( "4#浊环热水泵备妥" )
      Contact( "4#浊环热水电动蝶阀备妥" )
   END_RUNG wire#w1
   // the same network as SCL:
   #"4#浊环热水泵排气电磁阀"(READY := "4#浊环热水泵备妥" AND "4#浊环热水电动蝶阀备妥", OUT := "4#浊环热水泵排气电磁阀");   // "引水排气块"
END_REGION

REGION Network 33
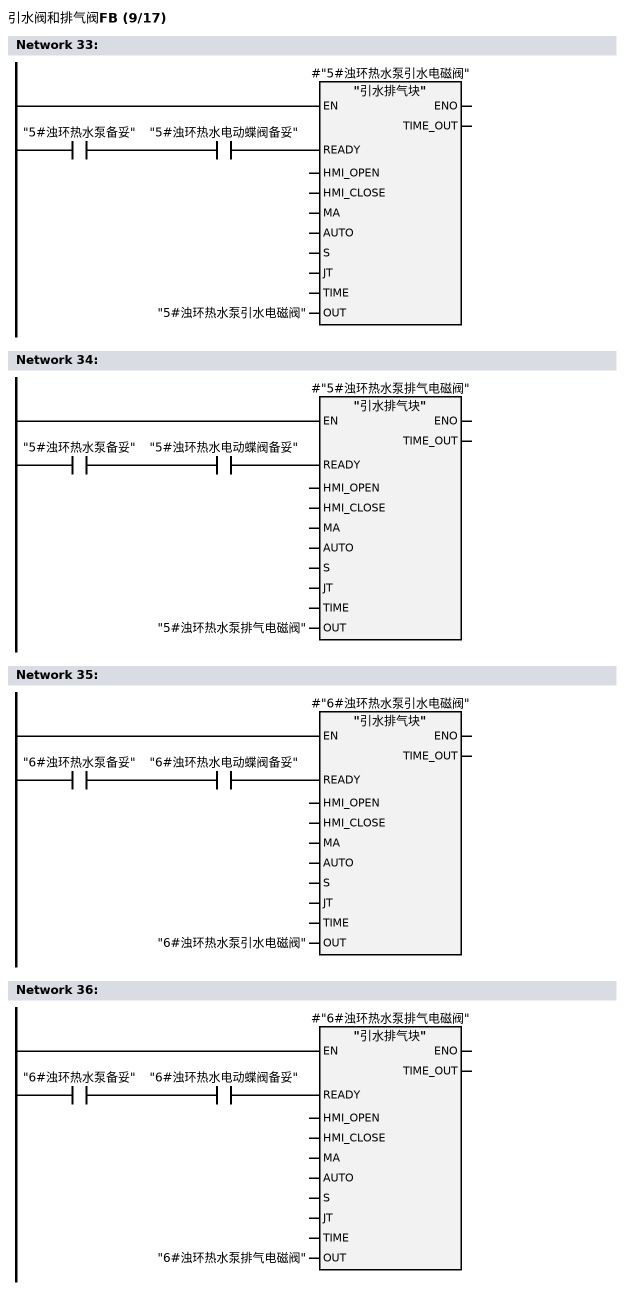
   RUNG wire#powerrail
      #"5#浊环热水泵引水电磁阀"(READY := wire#w1, HMI_OPEN :=, HMI_CLOSE :=, MA :=, AUTO :=, S :=, JT :=, "TIME" :=, OUT := "5#浊环热水泵引水电磁阀", TIME_OUT =>)
   END_RUNG
   RUNG wire#powerrail
      Contact( "5#浊环热水泵备妥" )
      Contact( "5#浊环热水电动蝶阀备妥" )
   END_RUNG wire#w1
   // the same network as SCL:
   #"5#浊环热水泵引水电磁阀"(READY := "5#浊环热水泵备妥" AND "5#浊环热水电动蝶阀备妥", OUT := "5#浊环热水泵引水电磁阀");   // "引水排气块"
END_REGION

REGION Network 34
   RUNG wire#powerrail
      #"5#浊环热水泵排气电磁阀"(READY := wire#w1, HMI_OPEN :=, HMI_CLOSE :=, MA :=, AUTO :=, S :=, JT :=, "TIME" :=, OUT := "5#浊环热水泵排气电磁阀", TIME_OUT =>)
   END_RUNG
   RUNG wire#powerrail
      Contact( "5#浊环热水泵备妥" )
      Contact( "5#浊环热水电动蝶阀备妥" )
   END_RUNG wire#w1
   // the same network as SCL:
   #"5#浊环热水泵排气电磁阀"(READY := "5#浊环热水泵备妥" AND "5#浊环热水电动蝶阀备妥", OUT := "5#浊环热水泵排气电磁阀");   // "引水排气块"
END_REGION

REGION Network 35
   RUNG wire#powerrail
      #"6#浊环热水泵引水电磁阀"(READY := wire#w1, HMI_OPEN :=, HMI_CLOSE :=, MA :=, AUTO :=, S :=, JT :=, "TIME" :=, OUT := "6#浊环热水泵引水电磁阀", TIME_OUT =>)
   END_RUNG
   RUNG wire#powerrail
      Contact( "6#浊环热水泵备妥" )
      Contact( "6#浊环热水电动蝶阀备妥" )
   END_RUNG wire#w1
   // the same network as SCL:
   #"6#浊环热水泵引水电磁阀"(READY := "6#浊环热水泵备妥" AND "6#浊环热水电动蝶阀备妥", OUT := "6#浊环热水泵引水电磁阀");   // "引水排气块"
END_REGION

REGION Network 36
   RUNG wire#powerrail
      #"6#浊环热水泵排气电磁阀"(READY := wire#w1, HMI_OPEN :=, HMI_CLOSE :=, MA :=, AUTO :=, S :=, JT :=, "TIME" :=, OUT := "6#浊环热水泵排气电磁阀", TIME_OUT =>)
   END_RUNG
   RUNG wire#powerrail
      Contact( "6#浊环热水泵备妥" )
      Contact( "6#浊环热水电动蝶阀备妥" )
   END_RUNG wire#w1
   // the same network as SCL:
   #"6#浊环热水泵排气电磁阀"(READY := "6#浊环热水泵备妥" AND "6#浊环热水电动蝶阀备妥", OUT := "6#浊环热水泵排气电磁阀");   // "引水排气块"
END_REGION

REGION Network 37
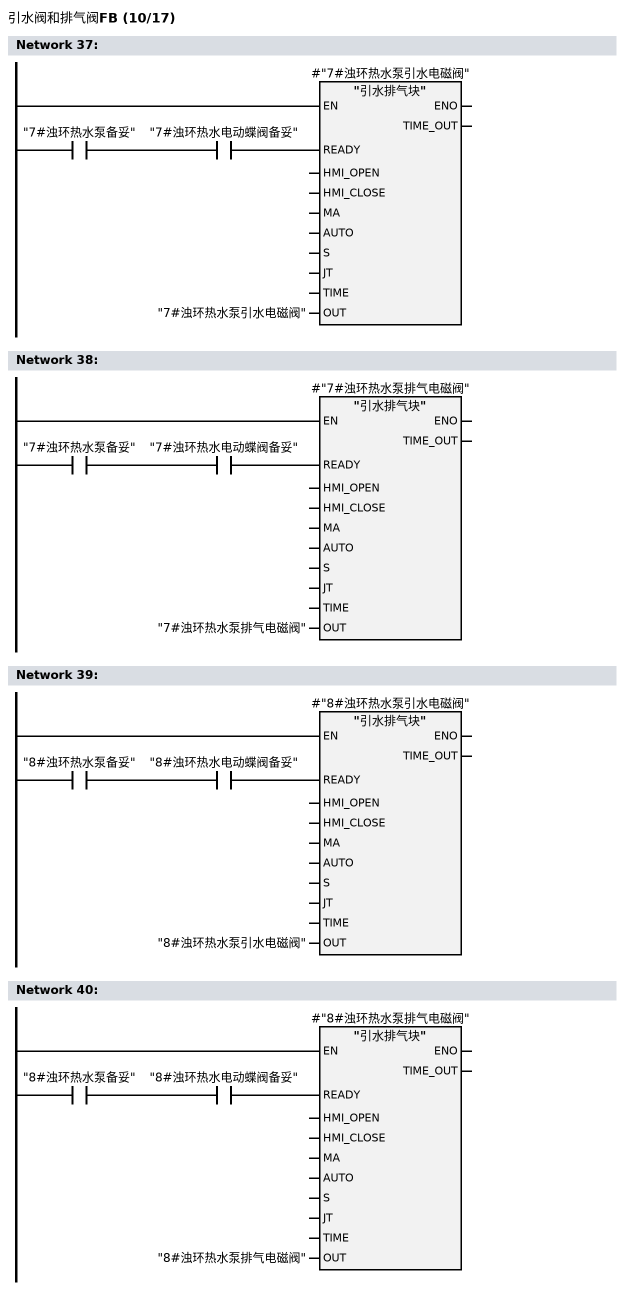
   RUNG wire#powerrail
      #"7#浊环热水泵引水电磁阀"(READY := wire#w1, HMI_OPEN :=, HMI_CLOSE :=, MA :=, AUTO :=, S :=, JT :=, "TIME" :=, OUT := "7#浊环热水泵引水电磁阀", TIME_OUT =>)
   END_RUNG
   RUNG wire#powerrail
      Contact( "7#浊环热水泵备妥" )
      Contact( "7#浊环热水电动蝶阀备妥" )
   END_RUNG wire#w1
   // the same network as SCL:
   #"7#浊环热水泵引水电磁阀"(READY := "7#浊环热水泵备妥" AND "7#浊环热水电动蝶阀备妥", OUT := "7#浊环热水泵引水电磁阀");   // "引水排气块"
END_REGION

REGION Network 38
   RUNG wire#powerrail
      #"7#浊环热水泵排气电磁阀"(READY := wire#w1, HMI_OPEN :=, HMI_CLOSE :=, MA :=, AUTO :=, S :=, JT :=, "TIME" :=, OUT := "7#浊环热水泵排气电磁阀", TIME_OUT =>)
   END_RUNG
   RUNG wire#powerrail
      Contact( "7#浊环热水泵备妥" )
      Contact( "7#浊环热水电动蝶阀备妥" )
   END_RUNG wire#w1
   // the same network as SCL:
   #"7#浊环热水泵排气电磁阀"(READY := "7#浊环热水泵备妥" AND "7#浊环热水电动蝶阀备妥", OUT := "7#浊环热水泵排气电磁阀");   // "引水排气块"
END_REGION
